REGION Network 3: Request Command
   RUNG wire#powerrail
      Contact( #Process.CmdRead )
      wire#w1
      I_Contact( #MB_CLIENT_Instance.BUSY )
      Coil( #MB_Ctrl.REQ )
   END_RUNG
   RUNG wire#powerrail
      Contact( #MB_Ctrl.REQ_Again )
   END_RUNG wire#w1
   // the same network as SCL:
   #MB_Ctrl.REQ := (#Process.CmdRead OR #MB_Ctrl.REQ_Again) AND NOT #MB_CLIENT_Instance.BUSY;
END_REGION

REGION Network 4: Retried Command
   #"Timer"."1".TON(IN := (#MB_CLIENT_Instance.ERROR OR (NOT #MB_CLIENT_Instance.ERROR AND NOT #MB_CLIENT_Instance.DONE)) AND NOT #MB_Ctrl.REQ_Again,
                    PT := T#5s);
   #MB_Ctrl.REQ_Again := #"Timer"."1".Q;
   #MB_CLIENT_Instance.Connected := #"Timer"."1".Q;
END_REGION

REGION Network 5: Modbus Client Instance call
   #MB_CLIENT_Instance(REQ := #MB_Ctrl.REQ,   // MB_CLIENT
                       DISCONNECT := #MB_Ctrl.Disconnect,
                       MB_MODE := #MB_Ctrl.MB_Mode,
                       MB_DATA_ADDR := #MB_Ctrl.MB_Data_Address,
                       MB_DATA_LEN := #MB_Ctrl.MB_Data_Length,
                       MB_DATA_PTR := #MB_Data.Buffer,
                       CONNECT := #MB_Ctrl.Connect);
END_REGION

REGION Network 6
   RUNG wire#powerrail
      Contact( #MB_CLIENT_Instance.BUSY )
      Coil( #Processing )
   END_RUNG
   RUNG wire#powerrail
      Contact( #MB_CLIENT_Instance.ERROR )
      Coil( #Error )
   END_RUNG
   // the same network as SCL:
   #Processing := #MB_CLIENT_Instance.BUSY;
   #Error := #MB_CLIENT_Instance.ERROR;
END_REGION
END_FUNCTION_BLOCK

FUNCTION_BLOCK "MFC_MB_iDT"   // FB27, LAD
TITLE = Modbus Block for Real Data Type
{ S7_Optimized_Access := 'TRUE' }
AUTHOR : JL
VERSION : 0.1
   VAR_INPUT
      InterfaceId : Hw_Any;   // HW-identifier of IE-interface submodule
      ID : Conn_Ouc;   // connection reference / identifier
      ConnectionType : Byte;   // type of connection: 11=TCP/IP, 19=UDP (17=TCP/IP)
      ActiveEstablished : Bool := true;   // active/passive connection establishment
      MB_Mode : Byte;
      ADDR1 : Byte;   // IPv4 address
      ADDR2 : Byte;   // IPv4 address
      ADDR3 : Byte;   // IPv4 address
      ADDR4 : Byte;   // IPv4 address
      RemotePort : UInt;   // remote UDP/TCP port number
      MB_Unit_ID : Byte;   // The Modbus slave address
      MB_Data_Add : UDInt;   // Modbus Data Address
      MB_Data_Len : UInt;   // Modbus Data Length
      FbkBusy : Bool;
      MultiFunction : Bool;   // Depend of the status of the other calls same MB
   END_VAR
   VAR_OUTPUT
      Busy : Bool;
      Done : Bool;
      Error : Bool;
      No_Connection : Bool;   // No connection with the Modbus Slave
      Status : Word;
   END_VAR
   VAR
      MB_CLIENT_Instance : MB_CLIENT;
      MB_Ctrl : Struct
         REQ : Bool;
         REQ_Again : Bool;
         Disconnect : Bool := false;
         MB_Mode : Byte;   // Modbus Mode
         MB_Data_Address : UDInt;   // Modbus Data Address
         MB_Data_Length : UInt;   // Modbus Data Length
         Connect : TCON_IP_v4;   // Connect Parameters Client
      END_STRUCT;
      MB_Data : Struct
         Buffer : Array[1..8] of Int;
      END_STRUCT;
      "Timer" : Struct
         "1" : IEC_TIMER;
         "2" : IEC_TIMER;
         ConnectionError : IEC_TIMER;
      END_STRUCT;
      OS : Struct
         bit : Array[0..31] of Bool;
      END_STRUCT;
      Process : Struct
         Start : Bool;
         CmdRead : Bool;
         End : Bool;
      END_STRUCT;
   END_VAR
   VAR_TEMP   // added for the SCL form of the ladder/FBD networks
      _w1 : Bool;
      _w2 : Bool;
      _w3 : Bool;
      _w4 : Bool;
   END_VAR
   // MB_Ctrl.Connect.InterfaceId := 258;
   // MB_Ctrl.Connect.ID := 11;
   // MB_Ctrl.Connect.ConnectionType := 11;
   // MB_Ctrl.Connect.ActiveEstablished := 1;
   // MB_Ctrl.Connect.RemoteAddress.ADDR[1] := 192;
   // MB_Ctrl.Connect.RemoteAddress.ADDR[2] := 168;
   // MB_Ctrl.Connect.RemoteAddress.ADDR[3] := 2;
   // MB_Ctrl.Connect.RemoteAddress.ADDR[4] := 11;
   // MB_Ctrl.Connect.RemotePort := 502;
BEGIN

REGION Network 1 (SCL): Block Parameters
   #MB_Ctrl.Connect.InterfaceId := #InterfaceId;
   #MB_Ctrl.Connect.ID := #ID;
   #MB_Ctrl.Connect.ConnectionType:=#ConnectionType;
   #MB_Ctrl.MB_Mode:=#MB_Mode;
   #MB_Ctrl.Connect.ActiveEstablished:=#ActiveEstablished;
   #MB_Ctrl.Connect.RemoteAddress.ADDR[1] := #ADDR1;
   #MB_Ctrl.Connect.RemoteAddress.ADDR[2] := #ADDR2;
   #MB_Ctrl.Connect.RemoteAddress.ADDR[3] := #ADDR3;
   #MB_Ctrl.Connect.RemoteAddress.ADDR[4] := #ADDR4;
   #MB_Ctrl.Connect.RemotePort := #RemotePort;
   #MB_CLIENT_Instance.MB_Unit_ID := #MB_Unit_ID;
   #MB_Ctrl.MB_Data_Address := #MB_Data_Add;
   #MB_Ctrl.MB_Data_Length := #MB_Data_Len;
   //#MB_Ctrl.Disconnect := #FbkBusy;
END_REGION

REGION Network 2: Reading Indication
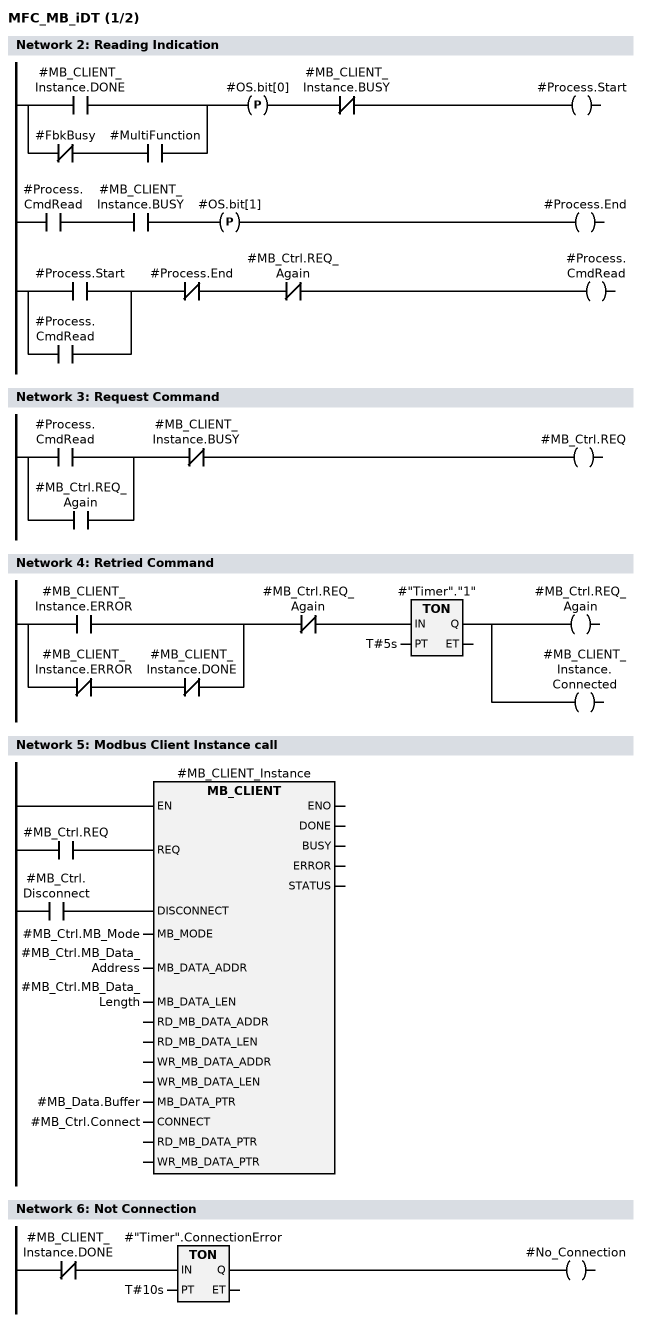
   RUNG wire#powerrail
      Contact( #MB_CLIENT_Instance.DONE )
      wire#w1
      P_Trig( #OS.bit[0] )
      I_Contact( #MB_CLIENT_Instance.BUSY )
      Coil( #Process.Start )
   END_RUNG
   RUNG wire#powerrail
      I_Contact( #FbkBusy )
      Contact( #MultiFunction )
   END_RUNG wire#w1
   RUNG wire#powerrail
      Contact( #Process.CmdRead )
      Contact( #MB_CLIENT_Instance.BUSY )
      P_Trig( #OS.bit[1] )
      Coil( #Process.End )
   END_RUNG
   RUNG wire#powerrail
      Contact( #Process.Start )
      wire#w2
      I_Contact( #Process.End )
      I_Contact( #MB_Ctrl.REQ_Again )
      Coil( #Process.CmdRead )
   END_RUNG
   RUNG wire#powerrail
      Contact( #Process.CmdRead )
   END_RUNG wire#w2
   // the same network as SCL:
   #_w1 := #MB_CLIENT_Instance.DONE OR (NOT #FbkBusy AND #MultiFunction);
   #_w2 := #_w1 AND NOT #OS.bit[0];   // rising edge
   #OS.bit[0] := #_w1;
   #Process.Start := #_w2 AND NOT #MB_CLIENT_Instance.BUSY;
   #_w3 := #Process.CmdRead AND #MB_CLIENT_Instance.BUSY;
   #_w4 := #_w3 AND NOT #OS.bit[1];   // rising edge
   #OS.bit[1] := #_w3;
   #Process.End := #_w4;
   #Process.CmdRead := (#Process.Start OR #Process.CmdRead) AND NOT #Process.End AND NOT #MB_Ctrl.REQ_Again;
END_REGION

REGION Network 3: Request Command
   RUNG wire#powerrail
      Contact( #Process.CmdRead )
      wire#w1
      I_Contact( #MB_CLIENT_Instance.BUSY )
      Coil( #MB_Ctrl.REQ )
   END_RUNG
   RUNG wire#powerrail
      Contact( #MB_Ctrl.REQ_Again )
   END_RUNG wire#w1
   // the same network as SCL:
   #MB_Ctrl.REQ := (#Process.CmdRead OR #MB_Ctrl.REQ_Again) AND NOT #MB_CLIENT_Instance.BUSY;
END_REGION

REGION Network 4: Retried Command
   #"Timer"."1".TON(IN := (#MB_CLIENT_Instance.ERROR OR (NOT #MB_CLIENT_Instance.ERROR AND NOT #MB_CLIENT_Instance.DONE)) AND NOT #MB_Ctrl.REQ_Again,
                    PT := T#5s);
   #MB_Ctrl.REQ_Again := #"Timer"."1".Q;
   #MB_CLIENT_Instance.Connected := #"Timer"."1".Q;
END_REGION

REGION Network 5: Modbus Client Instance call
   #MB_CLIENT_Instance(REQ := #MB_Ctrl.REQ,   // MB_CLIENT
                       DISCONNECT := #MB_Ctrl.Disconnect,
                       MB_MODE := #MB_Ctrl.MB_Mode,
                       MB_DATA_ADDR := #MB_Ctrl.MB_Data_Address,
                       MB_DATA_LEN := #MB_Ctrl.MB_Data_Length,
                       MB_DATA_PTR := #MB_Data.Buffer,
                       CONNECT := #MB_Ctrl.Connect);
END_REGION

REGION Network 6: Not Connection
   #"Timer".ConnectionError.TON(IN := NOT #MB_CLIENT_Instance.DONE, PT := T#10s);
   #No_Connection := #"Timer".ConnectionError.Q;
END_REGION

REGION Network 7: Block Status
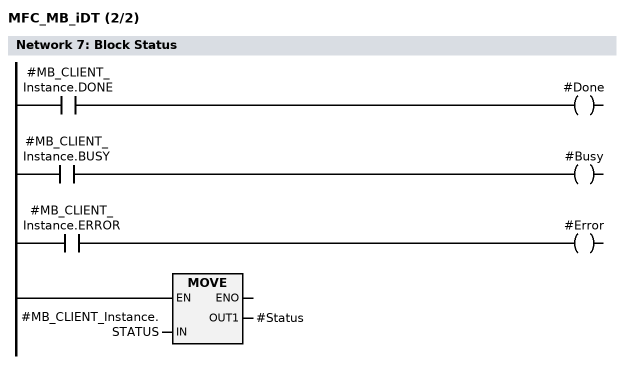
   RUNG wire#powerrail
      Contact( #MB_CLIENT_Instance.DONE )
      Coil( #Done )
   END_RUNG
   RUNG wire#powerrail
      Contact( #MB_CLIENT_Instance.BUSY )
      Coil( #Busy )
   END_RUNG
   RUNG wire#powerrail
      Contact( #MB_CLIENT_Instance.ERROR )
      Coil( #Error )
   END_RUNG
   RUNG wire#powerrail
      Move(in := #MB_CLIENT_Instance.STATUS, out1 => #Status)
   END_RUNG
   // the same network as SCL:
   #Done := #MB_CLIENT_Instance.DONE;
   #Busy := #MB_CLIENT_Instance.BUSY;
   #Error := #MB_CLIENT_Instance.ERROR;
   #Status := #MB_CLIENT_Instance.STATUS;
END_REGION
END_FUNCTION_BLOCK

FUNCTION_BLOCK "MFC_MB_ByteDT"   // FB35, LAD
TITLE = Modbus Block for Real Data Type
{ S7_Optimized_Access := 'TRUE' }
AUTHOR : JL
VERSION : 0.1
   VAR_INPUT
      InterfaceId : Hw_Any;   // HW-identifier of IE-interface submodule
      ID : Conn_Ouc;   // connection reference / identifier
      ConnectionType : Byte;   // type of connection: 11=TCP/IP, 19=UDP (17=TCP/IP)
      ActiveEstablished : Bool := true;   // active/passive connection establishment
      MB_Mode : Byte;
      ADDR1 : Byte;   // IPv4 address
      ADDR2 : Byte;   // IPv4 address
      ADDR3 : Byte;   // IPv4 address
      ADDR4 : Byte;   // IPv4 address
      RemotePort : UInt;   // remote UDP/TCP port number
      MB_Unit_ID : Byte;   // The Modbus slave address
      MB_Data_Add : UDInt;   // Modbus Data Address
      MB_Data_Len : UInt;   // Modbus Data Length
      FbkBusy : Bool;
      MultiFunction : Bool;   // Depend of the status of the other calls same MB
   END_VAR
   VAR_OUTPUT
      Busy : Bool;
      Done : Bool;
      Error : Bool;
      No_Connection : Bool;   // No connection with the Modbus Slave
      Status : Word;
   END_VAR
   VAR
      MB_CLIENT_Instance : MB_CLIENT;
      MB_Ctrl : Struct
         REQ : Bool;
         REQ_Again : Bool;
         Disconnect : Bool := false;
         MB_Mode : Byte;   // Modbus Mode
         MB_Data_Address : UDInt;   // Modbus Data Address
         MB_Data_Length : UInt;   // Modbus Data Length
         Connect : TCON_IP_v4;   // Connect Parameters Client
      END_STRUCT;
      MB_Data : Struct
         Buffer : Array[1..12] of Real;
      END_STRUCT;
      "Timer" : Struct
         "1" : IEC_TIMER;
         "2" : IEC_TIMER;
         ConnectionError : IEC_TIMER;
      END_STRUCT;
      OS : Struct
         bit : Array[0..31] of Bool;
      END_STRUCT;
      Process : Struct
         Start : Bool;
         CmdRead : Bool;
         End : Bool;
      END_STRUCT;
   END_VAR
   VAR_TEMP   // added for the SCL form of the ladder/FBD networks
      _w1 : Bool;
      _w2 : Bool;
      _w3 : Bool;
      _w4 : Bool;
   END_VAR
   // MB_Ctrl.Connect.InterfaceId := 258;
   // MB_Ctrl.Connect.ID := 11;
   // MB_Ctrl.Connect.ConnectionType := 11;
   // MB_Ctrl.Connect.ActiveEstablished := 1;
   // MB_Ctrl.Connect.RemoteAddress.ADDR[1] := 192;
   // MB_Ctrl.Connect.RemoteAddress.ADDR[2] := 168;
   // MB_Ctrl.Connect.RemoteAddress.ADDR[3] := 2;
   // MB_Ctrl.Connect.RemoteAddress.ADDR[4] := 11;
   // MB_Ctrl.Connect.RemotePort := 502;
BEGIN

REGION Network 1 (SCL): Block Parameters
   #MB_Ctrl.Connect.InterfaceId := #InterfaceId;
   #MB_Ctrl.Connect.ID := #ID;
   #MB_Ctrl.Connect.ConnectionType:=#ConnectionType;
   #MB_Ctrl.MB_Mode:=#MB_Mode;
   #MB_Ctrl.Connect.ActiveEstablished:=#ActiveEstablished;
   #MB_Ctrl.Connect.RemoteAddress.ADDR[1] := #ADDR1;
   #MB_Ctrl.Connect.RemoteAddress.ADDR[2] := #ADDR2;
   #MB_Ctrl.Connect.RemoteAddress.ADDR[3] := #ADDR3;
   #MB_Ctrl.Connect.RemoteAddress.ADDR[4] := #ADDR4;
   #MB_Ctrl.Connect.RemotePort := #RemotePort;
   #MB_CLIENT_Instance.MB_Unit_ID := #MB_Unit_ID;
   #MB_Ctrl.MB_Data_Address := #MB_Data_Add;
   #MB_Ctrl.MB_Data_Length := #MB_Data_Len;
   //#MB_Ctrl.Disconnect := #FbkBusy;
END_REGION

REGION Network 2: Reading Indication
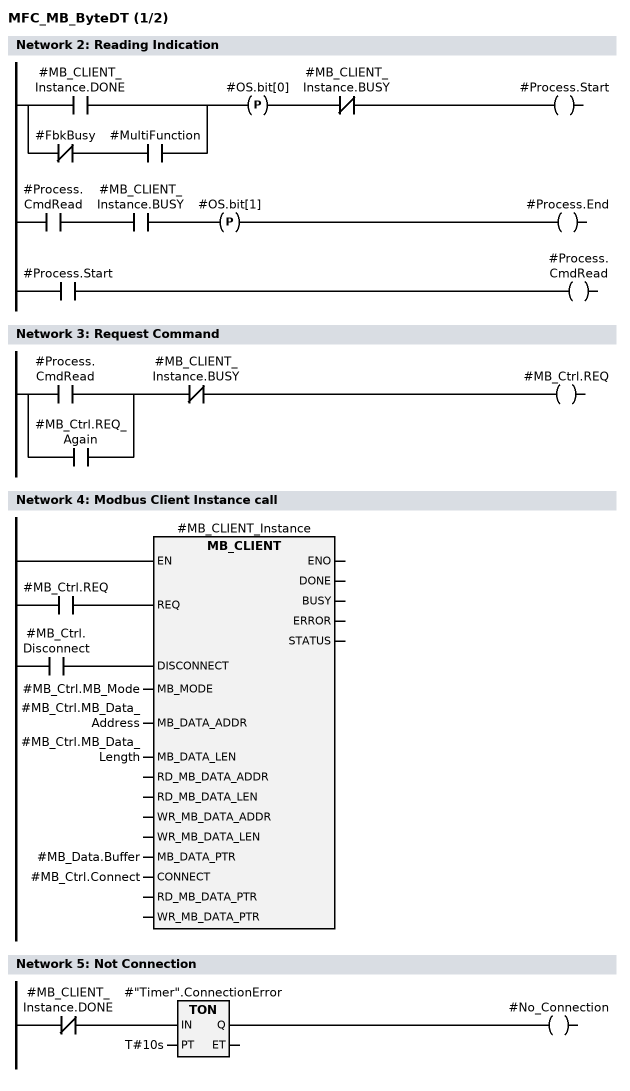
   RUNG wire#powerrail
      Contact( #MB_CLIENT_Instance.DONE )
      wire#w1
      P_Trig( #OS.bit[0] )
      I_Contact( #MB_CLIENT_Instance.BUSY )
      Coil( #Process.Start )
   END_RUNG
   RUNG wire#powerrail
      I_Contact( #FbkBusy )
      Contact( #MultiFunction )
   END_RUNG wire#w1
   RUNG wire#powerrail
      Contact( #Process.CmdRead )
      Contact( #MB_CLIENT_Instance.BUSY )
      P_Trig( #OS.bit[1] )
      Coil( #Process.End )
   END_RUNG
   RUNG wire#powerrail
      Contact( #Process.Start )
      Coil( #Process.CmdRead )
   END_RUNG
   // the same network as SCL:
   #_w1 := #MB_CLIENT_Instance.DONE OR (NOT #FbkBusy AND #MultiFunction);
   #_w2 := #_w1 AND NOT #OS.bit[0];   // rising edge
   #OS.bit[0] := #_w1;
   #Process.Start := #_w2 AND NOT #MB_CLIENT_Instance.BUSY;
   #_w3 := #Process.CmdRead AND #MB_CLIENT_Instance.BUSY;
   #_w4 := #_w3 AND NOT #OS.bit[1];   // rising edge
   #OS.bit[1] := #_w3;
   #Process.End := #_w4;
   #Process.CmdRead := #Process.Start;
END_REGION

REGION Network 3: Request Command
   RUNG wire#powerrail
      Contact( #Process.CmdRead )
      wire#w1
      I_Contact( #MB_CLIENT_Instance.BUSY )
      Coil( #MB_Ctrl.REQ )
   END_RUNG
   RUNG wire#powerrail
      Contact( #MB_Ctrl.REQ_Again )
   END_RUNG wire#w1
   // the same network as SCL:
   #MB_Ctrl.REQ := (#Process.CmdRead OR #MB_Ctrl.REQ_Again) AND NOT #MB_CLIENT_Instance.BUSY;
END_REGION

REGION Network 4: Modbus Client Instance call
   #MB_CLIENT_Instance(REQ := #MB_Ctrl.REQ,   // MB_CLIENT
                       DISCONNECT := #MB_Ctrl.Disconnect,
                       MB_MODE := #MB_Ctrl.MB_Mode,
                       MB_DATA_ADDR := #MB_Ctrl.MB_Data_Address,
                       MB_DATA_LEN := #MB_Ctrl.MB_Data_Length,
                       MB_DATA_PTR := #MB_Data.Buffer,
                       CONNECT := #MB_Ctrl.Connect);
END_REGION

REGION Network 5: Not Connection
   #"Timer".ConnectionError.TON(IN := NOT #MB_CLIENT_Instance.DONE, PT := T#10s);
   #No_Connection := #"Timer".ConnectionError.Q;
END_REGION

REGION Network 6: Block Status
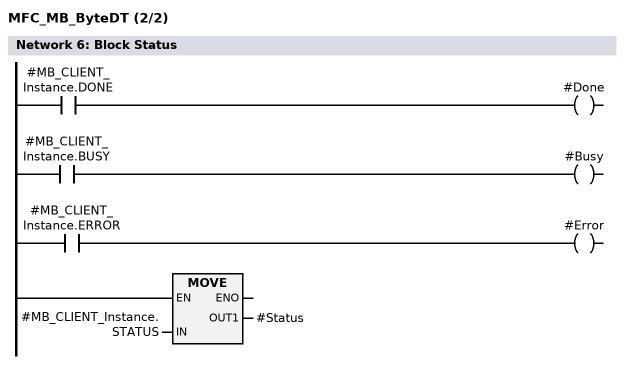
   RUNG wire#powerrail
      Contact( #MB_CLIENT_Instance.DONE )
      Coil( #Done )
   END_RUNG
   RUNG wire#powerrail
      Contact( #MB_CLIENT_Instance.BUSY )
      Coil( #Busy )
   END_RUNG
   RUNG wire#powerrail
      Contact( #MB_CLIENT_Instance.ERROR )
      Coil( #Error )
   END_RUNG
   RUNG wire#powerrail
      Move(in := #MB_CLIENT_Instance.STATUS, out1 => #Status)
   END_RUNG
   // the same network as SCL:
   #Done := #MB_CLIENT_Instance.DONE;
   #Busy := #MB_CLIENT_Instance.BUSY;
   #Error := #MB_CLIENT_Instance.ERROR;
   #Status := #MB_CLIENT_Instance.STATUS;
END_REGION
END_FUNCTION_BLOCK

// folder: Outside Comms/ModBus Comms/MFCs/MFC-4011

FUNCTION "MFC-4011_MB" : Void   // FC30, LAD
{ S7_Optimized_Access := 'TRUE' }
VERSION : 0.1
BEGIN

REGION Network 1: MFC Read Data Type Real
   // Read: 31203
   // *Pressure
   // *Flow Temperature
   // *Volumetric Flow
   // *Mass Flow
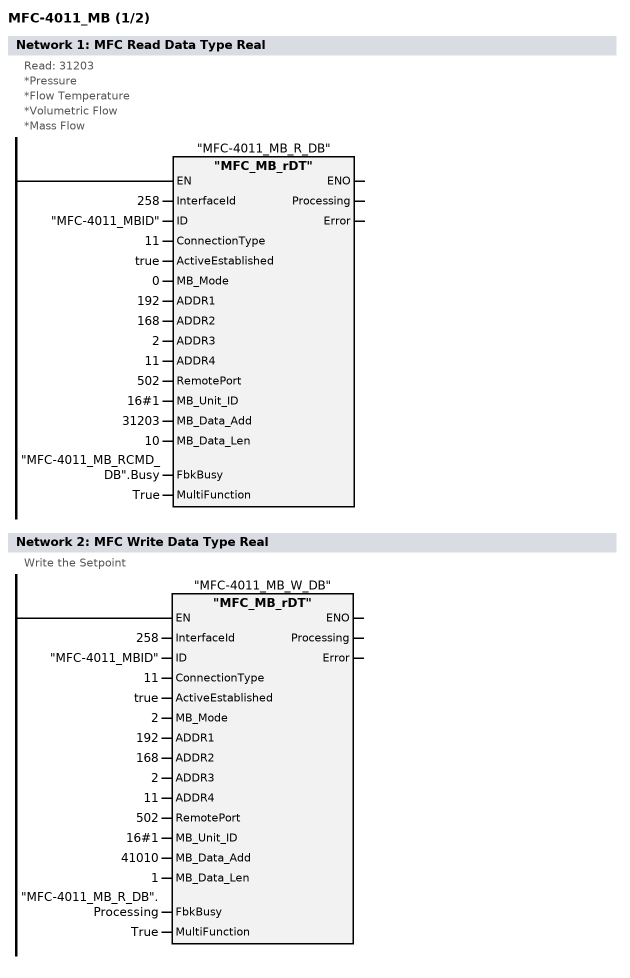
   RUNG wire#powerrail
      "MFC-4011_MB_R_DB"(InterfaceId := 258, ID := "MFC-4011_MBID", ConnectionType := 11, ActiveEstablished := true, MB_Mode := 0, ADDR1 := 192, ADDR2 := 168, ADDR3 := 2, ADDR4 := 11, RemotePort := 502, MB_Unit_ID := 16#1, MB_Data_Add := 31203, MB_Data_Len := 10, FbkBusy := "MFC-4011_MB_RCMD_DB".Busy, MultiFunction := True, Processing =>, Error =>)
   END_RUNG
   // the same network as SCL:
   "MFC-4011_MB_R_DB"(InterfaceId := 258,   // "MFC_MB_rDT"
                      ID := "MFC-4011_MBID",
                      ConnectionType := 11,
                      ActiveEstablished := true,
                      MB_Mode := 0,
                      ADDR1 := 192,
                      ADDR2 := 168,
                      ADDR3 := 2,
                      ADDR4 := 11,
                      RemotePort := 502,
                      MB_Unit_ID := 16#1,
                      MB_Data_Add := 31203,
                      MB_Data_Len := 10,
                      FbkBusy := "MFC-4011_MB_RCMD_DB".Busy,
                      MultiFunction := True);
END_REGION

REGION Network 2: MFC Write Data Type Real
   // Write the Setpoint
   RUNG wire#powerrail
      "MFC-4011_MB_W_DB"(InterfaceId := 258, ID := "MFC-4011_MBID", ConnectionType := 11, ActiveEstablished := true, MB_Mode := 2, ADDR1 := 192, ADDR2 := 168, ADDR3 := 2, ADDR4 := 11, RemotePort := 502, MB_Unit_ID := 16#1, MB_Data_Add := 41010, MB_Data_Len := 1, FbkBusy := "MFC-4011_MB_R_DB".Processing, MultiFunction := True, Processing =>, Error =>)
   END_RUNG
   // the same network as SCL:
   "MFC-4011_MB_W_DB"(InterfaceId := 258,   // "MFC_MB_rDT"
                      ID := "MFC-4011_MBID",
                      ConnectionType := 11,
                      ActiveEstablished := true,
                      MB_Mode := 2,
                      ADDR1 := 192,
                      ADDR2 := 168,
                      ADDR3 := 2,
                      ADDR4 := 11,
                      RemotePort := 502,
                      MB_Unit_ID := 16#1,
                      MB_Data_Add := 41010,
                      MB_Data_Len := 1,
                      FbkBusy := "MFC-4011_MB_R_DB".Processing,
                      MultiFunction := True);
END_REGION

REGION Network 3: MFC Write Data Type Int
   // Write the Command ID and the Command Argument
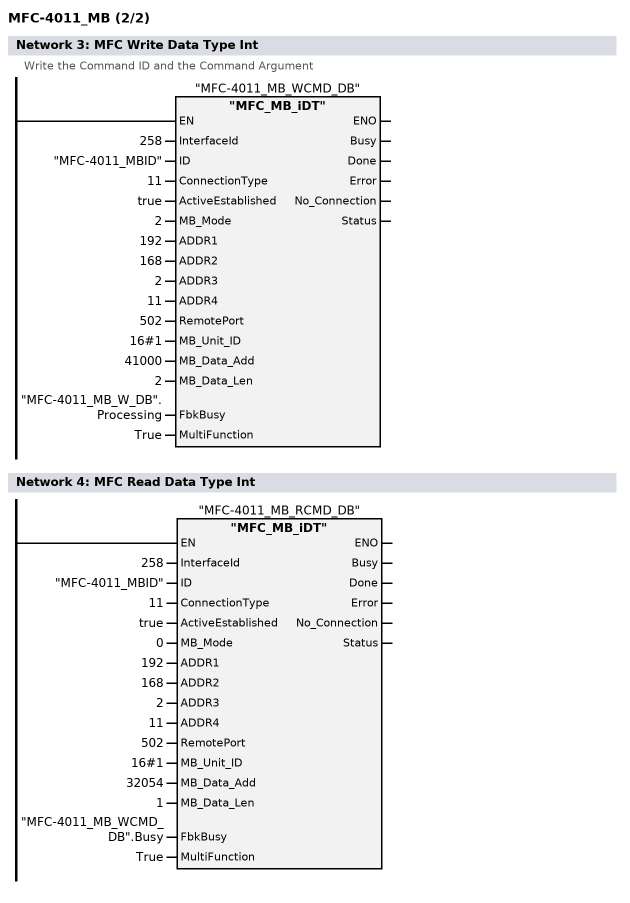
   RUNG wire#powerrail
      "MFC-4011_MB_WCMD_DB"(InterfaceId := 258, ID := "MFC-4011_MBID", ConnectionType := 11, ActiveEstablished := true, MB_Mode := 2, ADDR1 := 192, ADDR2 := 168, ADDR3 := 2, ADDR4 := 11, RemotePort := 502, MB_Unit_ID := 16#1, MB_Data_Add := 41000, MB_Data_Len := 2, FbkBusy := "MFC-4011_MB_W_DB".Processing, MultiFunction := True, Busy =>, Done =>, Error =>, No_Connection =>, Status =>)
   END_RUNG
   // the same network as SCL:
   "MFC-4011_MB_WCMD_DB"(InterfaceId := 258,   // "MFC_MB_iDT"
                         ID := "MFC-4011_MBID",
                         ConnectionType := 11,
                         ActiveEstablished := true,
                         MB_Mode := 2,
                         ADDR1 := 192,
                         ADDR2 := 168,
                         ADDR3 := 2,
                         ADDR4 := 11,
                         RemotePort := 502,
                         MB_Unit_ID := 16#1,
                         MB_Data_Add := 41000,
                         MB_Data_Len := 2,
                         FbkBusy := "MFC-4011_MB_W_DB".Processing,
                         MultiFunction := True);
END_REGION

REGION Network 4: MFC Read Data Type Int
   RUNG wire#powerrail
      "MFC-4011_MB_RCMD_DB"(InterfaceId := 258, ID := "MFC-4011_MBID", ConnectionType := 11, ActiveEstablished := true, MB_Mode := 0, ADDR1 := 192, ADDR2 := 168, ADDR3 := 2, ADDR4 := 11, RemotePort := 502, MB_Unit_ID := 16#1, MB_Data_Add := 32054, MB_Data_Len := 1, FbkBusy := "MFC-4011_MB_WCMD_DB".Busy, MultiFunction := True, Busy =>, Done =>, Error =>, No_Connection =>, Status =>)
   END_RUNG
   // the same network as SCL:
   "MFC-4011_MB_RCMD_DB"(InterfaceId := 258,   // "MFC_MB_iDT"
                         ID := "MFC-4011_MBID",
                         ConnectionType := 11,
                         ActiveEstablished := true,
                         MB_Mode := 0,
                         ADDR1 := 192,
                         ADDR2 := 168,
                         ADDR3 := 2,
                         ADDR4 := 11,
                         RemotePort := 502,
                         MB_Unit_ID := 16#1,
                         MB_Data_Add := 32054,
                         MB_Data_Len := 1,
                         FbkBusy := "MFC-4011_MB_WCMD_DB".Busy,
                         MultiFunction := True);
END_REGION
END_FUNCTION

// folder: Outside Comms/ModBus Comms/MFCs/MFC-4012

FUNCTION "MFC-4012_MB" : Void   // FC111, LAD
{ S7_Optimized_Access := 'TRUE' }
VERSION : 0.1
BEGIN

REGION Network 1: MFC Read Data Type Real
   // Read: 31203
   // *Pressure
   // *Flow Temperature
   // *Volumetric Flow
   // *Mass Flow
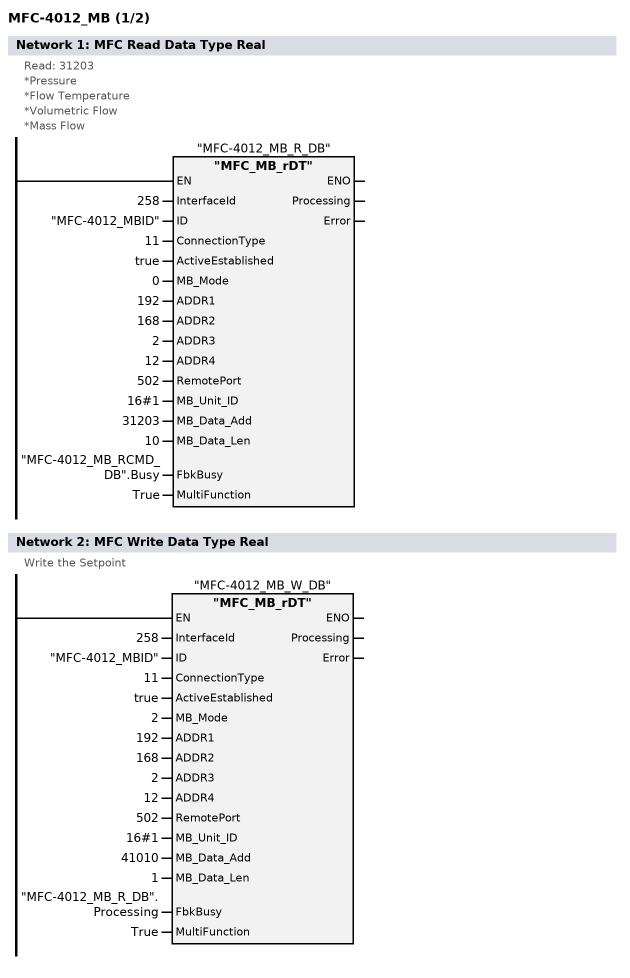
   RUNG wire#powerrail
      "MFC-4012_MB_R_DB"(InterfaceId := 258, ID := "MFC-4012_MBID", ConnectionType := 11, ActiveEstablished := true, MB_Mode := 0, ADDR1 := 192, ADDR2 := 168, ADDR3 := 2, ADDR4 := 12, RemotePort := 502, MB_Unit_ID := 16#1, MB_Data_Add := 31203, MB_Data_Len := 10, FbkBusy := "MFC-4012_MB_RCMD_DB".Busy, MultiFunction := True, Processing =>, Error =>)
   END_RUNG
   // the same network as SCL:
   "MFC-4012_MB_R_DB"(InterfaceId := 258,   // "MFC_MB_rDT"
                      ID := "MFC-4012_MBID",
                      ConnectionType := 11,
                      ActiveEstablished := true,
                      MB_Mode := 0,
                      ADDR1 := 192,
                      ADDR2 := 168,
                      ADDR3 := 2,
                      ADDR4 := 12,
                      RemotePort := 502,
                      MB_Unit_ID := 16#1,
                      MB_Data_Add := 31203,
                      MB_Data_Len := 10,
                      FbkBusy := "MFC-4012_MB_RCMD_DB".Busy,
                      MultiFunction := True);
END_REGION

REGION Network 2: MFC Write Data Type Real
   // Write the Setpoint
   RUNG wire#powerrail
      "MFC-4012_MB_W_DB"(InterfaceId := 258, ID := "MFC-4012_MBID", ConnectionType := 11, ActiveEstablished := true, MB_Mode := 2, ADDR1 := 192, ADDR2 := 168, ADDR3 := 2, ADDR4 := 12, RemotePort := 502, MB_Unit_ID := 16#1, MB_Data_Add := 41010, MB_Data_Len := 1, FbkBusy := "MFC-4012_MB_R_DB".Processing, MultiFunction := True, Processing =>, Error =>)
   END_RUNG
   // the same network as SCL:
   "MFC-4012_MB_W_DB"(InterfaceId := 258,   // "MFC_MB_rDT"
                      ID := "MFC-4012_MBID",
                      ConnectionType := 11,
                      ActiveEstablished := true,
                      MB_Mode := 2,
                      ADDR1 := 192,
                      ADDR2 := 168,
                      ADDR3 := 2,
                      ADDR4 := 12,
                      RemotePort := 502,
                      MB_Unit_ID := 16#1,
                      MB_Data_Add := 41010,
                      MB_Data_Len := 1,
                      FbkBusy := "MFC-4012_MB_R_DB".Processing,
                      MultiFunction := True);
END_REGION

REGION Network 3: MFC Write Data Type Int
   // Write the Command ID and the Command Argument
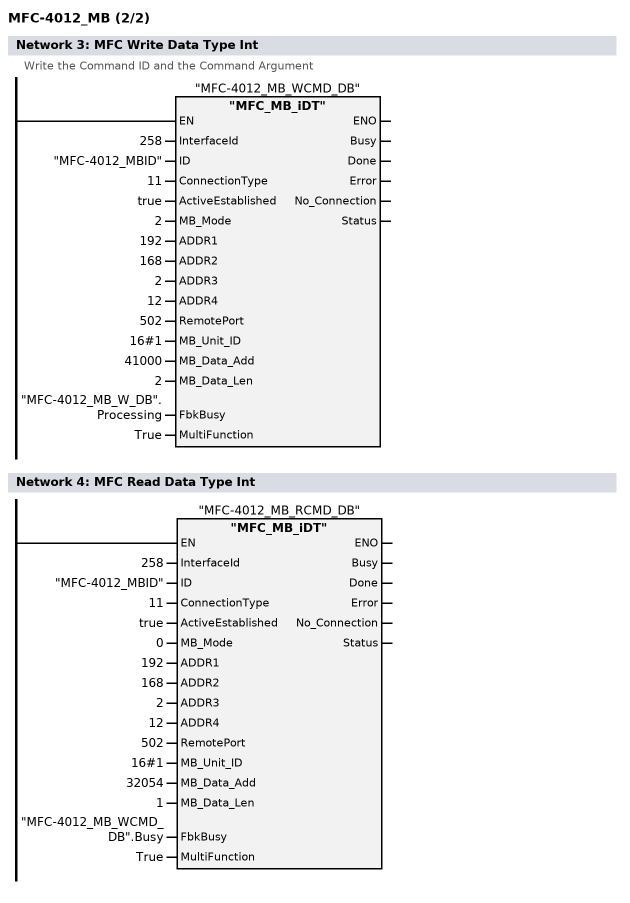
   RUNG wire#powerrail
      "MFC-4012_MB_WCMD_DB"(InterfaceId := 258, ID := "MFC-4012_MBID", ConnectionType := 11, ActiveEstablished := true, MB_Mode := 2, ADDR1 := 192, ADDR2 := 168, ADDR3 := 2, ADDR4 := 12, RemotePort := 502, MB_Unit_ID := 16#1, MB_Data_Add := 41000, MB_Data_Len := 2, FbkBusy := "MFC-4012_MB_W_DB".Processing, MultiFunction := True, Busy =>, Done =>, Error =>, No_Connection =>, Status =>)
   END_RUNG
   // the same network as SCL:
   "MFC-4012_MB_WCMD_DB"(InterfaceId := 258,   // "MFC_MB_iDT"
                         ID := "MFC-4012_MBID",
                         ConnectionType := 11,
                         ActiveEstablished := true,
                         MB_Mode := 2,
                         ADDR1 := 192,
                         ADDR2 := 168,
                         ADDR3 := 2,
                         ADDR4 := 12,
                         RemotePort := 502,
                         MB_Unit_ID := 16#1,
                         MB_Data_Add := 41000,
                         MB_Data_Len := 2,
                         FbkBusy := "MFC-4012_MB_W_DB".Processing,
                         MultiFunction := True);
END_REGION

REGION Network 4: MFC Read Data Type Int
   RUNG wire#powerrail
      "MFC-4012_MB_RCMD_DB"(InterfaceId := 258, ID := "MFC-4012_MBID", ConnectionType := 11, ActiveEstablished := true, MB_Mode := 0, ADDR1 := 192, ADDR2 := 168, ADDR3 := 2, ADDR4 := 12, RemotePort := 502, MB_Unit_ID := 16#1, MB_Data_Add := 32054, MB_Data_Len := 1, FbkBusy := "MFC-4012_MB_WCMD_DB".Busy, MultiFunction := True, Busy =>, Done =>, Error =>, No_Connection =>, Status =>)
   END_RUNG
   // the same network as SCL:
   "MFC-4012_MB_RCMD_DB"(InterfaceId := 258,   // "MFC_MB_iDT"
                         ID := "MFC-4012_MBID",
                         ConnectionType := 11,
                         ActiveEstablished := true,
                         MB_Mode := 0,
                         ADDR1 := 192,
                         ADDR2 := 168,
                         ADDR3 := 2,
                         ADDR4 := 12,
                         RemotePort := 502,
                         MB_Unit_ID := 16#1,
                         MB_Data_Add := 32054,
                         MB_Data_Len := 1,
                         FbkBusy := "MFC-4012_MB_WCMD_DB".Busy,
                         MultiFunction := True);
END_REGION
END_FUNCTION

// folder: Outside Comms/ModBus Comms/MFCs/MFC-4021

FUNCTION "MFC-4021_MB" : Void   // FC100, LAD
{ S7_Optimized_Access := 'TRUE' }
VERSION : 0.1
BEGIN

REGION Network 1: MFC Read Data Type Real
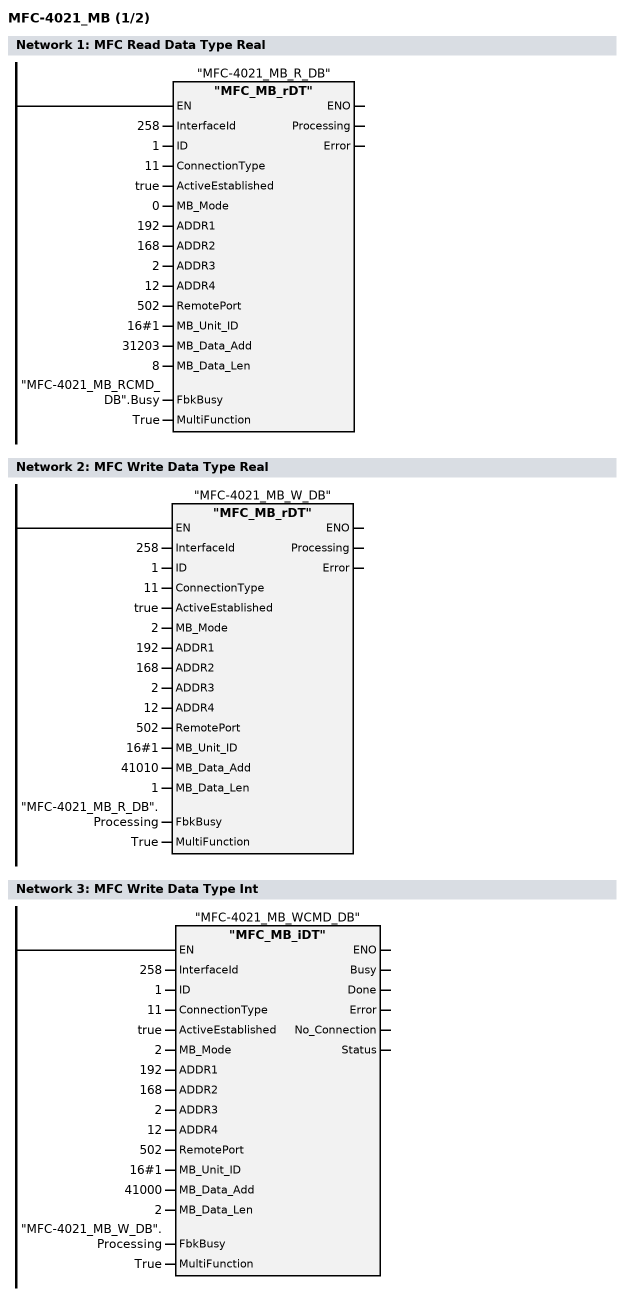
   RUNG wire#powerrail
      "MFC-4021_MB_R_DB"(InterfaceId := 258, ID := 1, ConnectionType := 11, ActiveEstablished := true, MB_Mode := 0, ADDR1 := 192, ADDR2 := 168, ADDR3 := 2, ADDR4 := 12, RemotePort := 502, MB_Unit_ID := 16#1, MB_Data_Add := 31203, MB_Data_Len := 8, FbkBusy := "MFC-4021_MB_RCMD_DB".Busy, MultiFunction := True, Processing =>, Error =>)
   END_RUNG
   // the same network as SCL:
   "MFC-4021_MB_R_DB"(InterfaceId := 258,   // "MFC_MB_rDT"
                      ID := 1,
                      ConnectionType := 11,
                      ActiveEstablished := true,
                      MB_Mode := 0,
                      ADDR1 := 192,
                      ADDR2 := 168,
                      ADDR3 := 2,
                      ADDR4 := 12,
                      RemotePort := 502,
                      MB_Unit_ID := 16#1,
                      MB_Data_Add := 31203,
                      MB_Data_Len := 8,
                      FbkBusy := "MFC-4021_MB_RCMD_DB".Busy,
                      MultiFunction := True);
END_REGION

REGION Network 2: MFC Write Data Type Real
   RUNG wire#powerrail
      "MFC-4021_MB_W_DB"(InterfaceId := 258, ID := 1, ConnectionType := 11, ActiveEstablished := true, MB_Mode := 2, ADDR1 := 192, ADDR2 := 168, ADDR3 := 2, ADDR4 := 12, RemotePort := 502, MB_Unit_ID := 16#1, MB_Data_Add := 41010, MB_Data_Len := 1, FbkBusy := "MFC-4021_MB_R_DB".Processing, MultiFunction := True, Processing =>, Error =>)
   END_RUNG
   // the same network as SCL:
   "MFC-4021_MB_W_DB"(InterfaceId := 258,   // "MFC_MB_rDT"
                      ID := 1,
                      ConnectionType := 11,
                      ActiveEstablished := true,
                      MB_Mode := 2,
                      ADDR1 := 192,
                      ADDR2 := 168,
                      ADDR3 := 2,
                      ADDR4 := 12,
                      RemotePort := 502,
                      MB_Unit_ID := 16#1,
                      MB_Data_Add := 41010,
                      MB_Data_Len := 1,
                      FbkBusy := "MFC-4021_MB_R_DB".Processing,
                      MultiFunction := True);
END_REGION

REGION Network 3: MFC Write Data Type Int
   RUNG wire#powerrail
      "MFC-4021_MB_WCMD_DB"(InterfaceId := 258, ID := 1, ConnectionType := 11, ActiveEstablished := true, MB_Mode := 2, ADDR1 := 192, ADDR2 := 168, ADDR3 := 2, ADDR4 := 12, RemotePort := 502, MB_Unit_ID := 16#1, MB_Data_Add := 41000, MB_Data_Len := 2, FbkBusy := "MFC-4021_MB_W_DB".Processing, MultiFunction := True, Busy =>, Done =>, Error =>, No_Connection =>, Status =>)
   END_RUNG
   // the same network as SCL:
   "MFC-4021_MB_WCMD_DB"(InterfaceId := 258,   // "MFC_MB_iDT"
                         ID := 1,
                         ConnectionType := 11,
                         ActiveEstablished := true,
                         MB_Mode := 2,
                         ADDR1 := 192,
                         ADDR2 := 168,
                         ADDR3 := 2,
                         ADDR4 := 12,
                         RemotePort := 502,
                         MB_Unit_ID := 16#1,
                         MB_Data_Add := 41000,
                         MB_Data_Len := 2,
                         FbkBusy := "MFC-4021_MB_W_DB".Processing,
                         MultiFunction := True);
END_REGION

REGION Network 4: MFC Read Data Type Int
